
ScreenModuleEditorView "Settings Station Row" 671x200
   TextField "tfLine" at 0,0 size 215x200; Text '$T'
      Visibility <- "Interface.line.visibility"
      Appearance <- "Interface.line.animate"
   TextField "tfLablBtn00" at 215,0 size 40x25; Text '1'
      Visibility <- "Interface.btnRows[0].button.visibility"
      Appearance <- "Interface.btnRows[0].button.animate"
   TextField "tfAllottedBtn00" at 255,0 size 80x25; Text 'Text'
      Visibility <- "Interface.btnRows[0].total.visibility"
      Appearance <- "Interface.btnRows[0].total.animate"
   TextField "tfCriticalBtn00" at 335,0 size 80x25; Text 'Text'
      Visibility <- "Interface.btnRows[0].critical.visibility"
      Appearance <- "Interface.btnRows[0].critical.animate"
   TextField "tfPartNumberBtn00" at 415,0 size 256x25; Text 'Text'
      Visibility <- "Interface.btnRows[0].singlePN.visibility"
      Appearance <- "Interface.btnRows[0].singlePN.animate"
   TextField "tfLablBtn01" at 215,25 size 40x25; Text '2'
      Visibility <- "Interface.btnRows[1].button.visibility"
      Appearance <- "Interface.btnRows[1].button.animate"
   TextField "tfAllottedBtn01" at 255,25 size 80x25; Text 'Text'
      Visibility <- "Interface.btnRows[1].total.visibility"
      Appearance <- "Interface.btnRows[1].total.animate"
   TextField "tfCriticalBtn01" at 335,25 size 80x25; Text 'Text'
      Visibility <- "Interface.btnRows[1].critical.visibility"
      Appearance <- "Interface.btnRows[1].critical.animate"
   TextField "tfPartNumberBtn01" at 415,25 size 256x25; Text 'Text'
      Visibility <- "Interface.btnRows[1].singlePN.visibility"
      Appearance <- "Interface.btnRows[1].singlePN.animate"
   TextField "tfLablBtn02" at 215,50 size 40x25; Text '3'
      Visibility <- "Interface.btnRows[2].button.visibility"
      Appearance <- "Interface.btnRows[2].button.animate"
   TextField "tfAllottedBtn02" at 255,50 size 80x25; Text 'Text'
      Visibility <- "Interface.btnRows[2].total.visibility"
      Appearance <- "Interface.btnRows[2].total.animate"
   TextField "tfCriticalBtn02" at 335,50 size 80x25; Text 'Text'
      Visibility <- "Interface.btnRows[2].critical.visibility"
      Appearance <- "Interface.btnRows[2].critical.animate"
   TextField "tfPartNumberBtn02" at 415,50 size 256x25; Text 'Text'
      Visibility <- "Interface.btnRows[2].singlePN.visibility"
      Appearance <- "Interface.btnRows[2].singlePN.animate"
   TextField "tfLablBtn03" at 215,75 size 40x25; Text '4'
      Visibility <- "Interface.btnRows[3].button.visibility"
      Appearance <- "Interface.btnRows[3].button.animate"
   TextField "tfAllottedBtn03" at 255,75 size 80x25; Text 'Text'
      Visibility <- "Interface.btnRows[3].total.visibility"
      Appearance <- "Interface.btnRows[3].total.animate"
   TextField "tfCriticalBtn03" at 335,75 size 80x25; Text 'Text'
      Visibility <- "Interface.btnRows[3].critical.visibility"
      Appearance <- "Interface.btnRows[3].critical.animate"
   TextField "tfPartNumberBtn03" at 415,75 size 256x25; Text 'Text'
      Visibility <- "Interface.btnRows[3].singlePN.visibility"
      Appearance <- "Interface.btnRows[3].singlePN.animate"
   TextField "tfLablBtn04" at 215,100 size 40x25; Text '5'
      Visibility <- "Interface.btnRows[4].button.visibility"
      Appearance <- "Interface.btnRows[4].button.animate"
   TextField "tfAllottedBtn04" at 255,100 size 80x25; Text 'Text'
      Visibility <- "Interface.btnRows[4].total.visibility"
      Appearance <- "Interface.btnRows[4].total.animate"
   TextField "tfCriticalBtn04" at 335,100 size 80x25; Text 'Text'
      Visibility <- "Interface.btnRows[4].critical.visibility"
      Appearance <- "Interface.btnRows[4].critical.animate"
   TextField "tfPartNumberBtn04" at 415,100 size 256x25; Text 'Text'
      Visibility <- "Interface.btnRows[4].singlePN.visibility"
      Appearance <- "Interface.btnRows[4].singlePN.animate"
   TextField "tfLablBtn05" at 215,125 size 40x25; Text '6'
      Visibility <- "Interface.btnRows[5].button.visibility"
      Appearance <- "Interface.btnRows[5].button.animate"
   TextField "tfAllottedBtn05" at 255,125 size 80x25; Text 'Text'
      Visibility <- "Interface.btnRows[5].total.visibility"
      Appearance <- "Interface.btnRows[5].total.animate"
   TextField "tfCriticalBtn05" at 335,125 size 80x25; Text 'Text'
      Visibility <- "Interface.btnRows[5].critical.visibility"
      Appearance <- "Interface.btnRows[5].critical.animate"
   TextField "tfPartNumberBtn05" at 415,125 size 256x25; Text 'Text'
      Visibility <- "Interface.btnRows[5].singlePN.visibility"
      Appearance <- "Interface.btnRows[5].singlePN.animate"
   TextField "tfLablBtn06" at 215,150 size 40x25; Text '7'
      Visibility <- "Interface.btnRows[6].button.visibility"
      Appearance <- "Interface.btnRows[6].button.animate"
   TextField "tfAllottedBtn06" at 255,150 size 80x25; Text 'Text'
      Visibility <- "Interface.btnRows[6].total.visibility"
      Appearance <- "Interface.btnRows[6].total.animate"
   TextField "tfCriticalBtn06" at 335,150 size 80x25; Text 'Text'
      Visibility <- "Interface.btnRows[6].critical.visibility"
      Appearance <- "Interface.btnRows[6].critical.animate"
   TextField "tfPartNumberBtn06" at 415,150 size 256x25; Text 'Text'
      Visibility <- "Interface.btnRows[6].singlePN.visibility"
      Appearance <- "Interface.btnRows[6].singlePN.animate"
   TextField "tfLablBtn07" at 215,175 size 40x25; Text '8'
      Visibility <- "Interface.btnRows[7].button.visibility"
      Appearance <- "Interface.btnRows[7].button.animate"
   TextField "tfAllottedBtn07" at 255,175 size 80x25; Text 'Text'
      Visibility <- "Interface.btnRows[7].total.visibility"
      Appearance <- "Interface.btnRows[7].total.animate"
   TextField "tfCriticalBtn07" at 335,175 size 80x25; Text 'Text'
      Visibility <- "Interface.btnRows[7].critical.visibility"
      Appearance <- "Interface.btnRows[7].critical.animate"
   TextField "tfPartNumberBtn07" at 415,175 size 256x25; Text 'Text'
      Visibility <- "Interface.btnRows[7].singlePN.visibility"
      Appearance <- "Interface.btnRows[7].singlePN.animate"
   TextField "tfPNDoubleBtn00" at 415,0 size 256x25; Text 'Text'
      Visibility <- "Interface.btnRows[0].doublePN.visibility"
      Appearance <- "Interface.btnRows[0].doublePN.animate"
   TextField "tfPNDoubleBtn01" at 415,25 size 256x25; Text 'Text'
      Visibility <- "Interface.btnRows[1].doublePN.visibility"
      Appearance <- "Interface.btnRows[1].doublePN.animate"
   TextField "tfPNDoubleBtn02" at 415,50 size 256x25; Text 'Text'
      Visibility <- "Interface.btnRows[2].doublePN.visibility"
      Appearance <- "Interface.btnRows[2].doublePN.animate"
   TextField "tfPNDoubleBtn03" at 415,75 size 256x25; Text 'Text'
      Visibility <- "Interface.btnRows[3].doublePN.visibility"
      Appearance <- "Interface.btnRows[3].doublePN.animate"
   TextField "tfPNDoubleBtn04" at 415,100 size 256x25; Text 'Text'
      Visibility <- "Interface.btnRows[4].doublePN.visibility"
      Appearance <- "Interface.btnRows[4].doublePN.animate"
   TextField "tfPNDoubleBtn05" at 415,125 size 256x25; Text 'Text'
      Visibility <- "Interface.btnRows[5].doublePN.visibility"
      Appearance <- "Interface.btnRows[5].doublePN.animate"
   TextField "tfPNDoubleBtn06" at 415,150 size 256x25; Text 'Text'
      Visibility <- "Interface.btnRows[6].doublePN.visibility"
      Appearance <- "Interface.btnRows[6].doublePN.animate"
   TextField "tfPNDoubleBtn07" at 415,175 size 256x25; Text 'Text'
      Visibility <- "Interface.btnRows[7].doublePN.visibility"
      Appearance <- "Interface.btnRows[7].doublePN.animate"
*)

(* ===== HMI "HMI_RT_1" =====

ScreenModuleEditorView "Settings Station Row" 671x200
   TextField "tfLine" at 0,0 size 215x200; Text 'Text'
      Visibility <- "Interface.line.visibility"
      Appearance <- "Interface.line.animate"
   TextField "tfLablBtn00" at 215,0 size 40x25; Text '1'
      Visibility <- "Interface.btnRows[0].button.visibility"
      Appearance <- "Interface.btnRows[0].button.animate"
   TextField "tfAllottedBtn00" at 255,0 size 80x25; Text 'Text'
      Visibility <- "Interface.btnRows[0].total.visibility"
      Appearance <- "Interface.btnRows[0].total.animate"
   TextField "tfCriticalBtn00" at 335,0 size 80x25; Text 'Text'
      Visibility <- "Interface.btnRows[0].critical.visibility"
      Appearance <- "Interface.btnRows[0].critical.animate"
   TextField "tfPartNumberBtn00" at 415,0 size 256x25; Text 'Text'
      Visibility <- "Interface.btnRows[0].singlePN.visibility"
      Appearance <- "Interface.btnRows[0].singlePN.animate"
   TextField "tfLablBtn01" at 215,25 size 40x25; Text '2'
      Visibility <- "Interface.btnRows[1].button.visibility"
      Appearance <- "Interface.btnRows[1].button.animate"
   TextField "tfAllottedBtn01" at 255,25 size 80x25; Text 'Text'
      Visibility <- "Interface.btnRows[1].total.visibility"
      Appearance <- "Interface.btnRows[1].total.animate"
   TextField "tfCriticalBtn01" at 335,25 size 80x25; Text 'Text'
      Visibility <- "Interface.btnRows[1].critical.visibility"
      Appearance <- "Interface.btnRows[1].critical.animate"
   TextField "tfPartNumberBtn01" at 415,25 size 256x25; Text 'Text'
      Visibility <- "Interface.btnRows[1].singlePN.visibility"
      Appearance <- "Interface.btnRows[1].singlePN.animate"
   TextField "tfLablBtn02" at 215,50 size 40x25; Text '3'
      Visibility <- "Interface.btnRows[2].button.visibility"
      Appearance <- "Interface.btnRows[2].button.animate"
   TextField "tfAllottedBtn02" at 255,50 size 80x25; Text 'Text'
      Visibility <- "Interface.btnRows[2].total.visibility"
      Appearance <- "Interface.btnRows[2].total.animate"
   TextField "tfCriticalBtn02" at 335,50 size 80x25; Text 'Text'
      Visibility <- "Interface.btnRows[2].critical.visibility"
      Appearance <- "Interface.btnRows[2].critical.animate"
   TextField "tfPartNumberBtn02" at 415,50 size 256x25; Text 'Text'
      Visibility <- "Interface.btnRows[2].singlePN.visibility"
      Appearance <- "Interface.btnRows[2].singlePN.animate"
   TextField "tfLablBtn03" at 215,75 size 40x25; Text '4'
      Visibility <- "Interface.btnRows[3].button.visibility"
      Appearance <- "Interface.btnRows[3].button.animate"
   TextField "tfAllottedBtn03" at 255,75 size 80x25; Text 'Text'
      Visibility <- "Interface.btnRows[3].total.visibility"
      Appearance <- "Interface.btnRows[3].total.animate"
   TextField "tfCriticalBtn03" at 335,75 size 80x25; Text 'Text'
      Visibility <- "Interface.btnRows[3].critical.visibility"
      Appearance <- "Interface.btnRows[3].critical.animate"
   TextField "tfPartNumberBtn03" at 415,75 size 256x25; Text 'Text'
      Visibility <- "Interface.btnRows[3].singlePN.visibility"
      Appearance <- "Interface.btnRows[3].singlePN.animate"
   TextField "tfLablBtn04" at 215,100 size 40x25; Text '5'
      Visibility <- "Interface.btnRows[4].button.visibility"
      Appearance <- "Interface.btnRows[4].button.animate"
   TextField "tfAllottedBtn04" at 255,100 size 80x25; Text 'Text'
      Visibility <- "Interface.btnRows[4].total.visibility"
      Appearance <- "Interface.btnRows[4].total.animate"
   TextField "tfCriticalBtn04" at 335,100 size 80x25; Text 'Text'
      Visibility <- "Interface.btnRows[4].critical.visibility"
      Appearance <- "Interface.btnRows[4].critical.animate"
   TextField "tfPartNumberBtn04" at 415,100 size 256x25; Text 'Text'
      Visibility <- "Interface.btnRows[4].singlePN.visibility"
      Appearance <- "Interface.btnRows[4].singlePN.animate"
   TextField "tfLablBtn05" at 215,125 size 40x25; Text '6'
      Visibility <- "Interface.btnRows[5].button.visibility"
      Appearance <- "Interface.btnRows[5].button.animate"
   TextField "tfAllottedBtn05" at 255,125 size 80x25; Text 'Text'
      Visibility <- "Interface.btnRows[5].total.visibility"
      Appearance <- "Interface.btnRows[5].total.animate"
   TextField "tfCriticalBtn05" at 335,125 size 80x25; Text 'Text'
      Visibility <- "Interface.btnRows[5].critical.visibility"
      Appearance <- "Interface.btnRows[5].critical.animate"
   TextField "tfPartNumberBtn05" at 415,125 size 256x25; Text 'Text'
      Visibility <- "Interface.btnRows[5].singlePN.visibility"
      Appearance <- "Interface.btnRows[5].singlePN.animate"
   TextField "tfLablBtn06" at 215,150 size 40x25; Text '7'
      Visibility <- "Interface.btnRows[6].button.visibility"
      Appearance <- "Interface.btnRows[6].button.animate"
   TextField "tfAllottedBtn06" at 255,150 size 80x25; Text 'Text'
      Visibility <- "Interface.btnRows[6].total.visibility"
      Appearance <- "Interface.btnRows[6].total.animate"
   TextField "tfCriticalBtn06" at 335,150 size 80x25; Text 'Text'
      Visibility <- "Interface.btnRows[6].critical.visibility"
      Appearance <- "Interface.btnRows[6].critical.animate"
   TextField "tfPartNumberBtn06" at 415,150 size 256x25; Text 'Text'
      Visibility <- "Interface.btnRows[6].singlePN.visibility"
      Appearance <- "Interface.btnRows[6].singlePN.animate"
   TextField "tfLablBtn07" at 215,175 size 40x25; Text '8'
      Visibility <- "Interface.btnRows[7].button.visibility"
      Appearance <- "Interface.btnRows[7].button.animate"
   TextField "tfAllottedBtn07" at 255,175 size 80x25; Text 'Text'
      Visibility <- "Interface.btnRows[7].total.visibility"
      Appearance <- "Interface.btnRows[7].total.animate"
   TextField "tfCriticalBtn07" at 335,175 size 80x25; Text 'Text'
      Visibility <- "Interface.btnRows[7].critical.visibility"
      Appearance <- "Interface.btnRows[7].critical.animate"
   TextField "tfPartNumberBtn07" at 415,175 size 256x25; Text 'Text'
      Visibility <- "Interface.btnRows[7].singlePN.visibility"
      Appearance <- "Interface.btnRows[7].singlePN.animate"
   TextField "tfPNDoubleBtn00" at 415,0 size 256x25; Text 'Text'
      Visibility <- "Interface.btnRows[0].doublePN.visibility"
      Appearance <- "Interface.btnRows[0].doublePN.animate"
   TextField "tfPNDoubleBtn01" at 415,25 size 256x25; Text 'Text'
      Visibility <- "Interface.btnRows[1].doublePN.visibility"
      Appearance <- "Interface.btnRows[1].doublePN.animate"
   TextField "tfPNDoubleBtn02" at 415,50 size 256x25; Text 'Text'
      Visibility <- "Interface.btnRows[2].doublePN.visibility"
      Appearance <- "Interface.btnRows[2].doublePN.animate"
   TextField "tfPNDoubleBtn03" at 415,75 size 256x25; Text 'Text'
      Visibility <- "Interface.btnRows[3].doublePN.visibility"
      Appearance <- "Interface.btnRows[3].doublePN.animate"
   TextField "tfPNDoubleBtn04" at 415,100 size 256x25; Text 'Text'
      Visibility <- "Interface.btnRows[4].doublePN.visibility"
      Appearance <- "Interface.btnRows[4].doublePN.animate"
   TextField "tfPNDoubleBtn05" at 415,125 size 256x25; Text 'Text'
      Visibility <- "Interface.btnRows[5].doublePN.visibility"
      Appearance <- "Interface.btnRows[5].doublePN.animate"
   TextField "tfPNDoubleBtn06" at 415,150 size 256x25; Text 'Text'
      Visibility <- "Interface.btnRows[6].doublePN.visibility"
      Appearance <- "Interface.btnRows[6].doublePN.animate"
   TextField "tfPNDoubleBtn07" at 415,175 size 256x25; Text 'Text'
      Visibility <- "Interface.btnRows[7].doublePN.visibility"
      Appearance <- "Interface.btnRows[7].doublePN.animate"
*)

(* ===== HMI "HMI_RT_1" =====

ScreenModuleEditorView "Settings Station Row" 671x200
   TextField "tfLine" at 0,0 size 215x200; Text 'Text'
      Visibility <- "Interface.line.visibility"
      Appearance <- "Interface.line.animate"
   TextField "tfLablBtn00" at 215,0 size 40x25; Text '1'
      Visibility <- "Interface.btnRows[0].button.visibility"
      Appearance <- "Interface.btnRows[0].button.animate"
   TextField "tfAllottedBtn00" at 255,0 size 80x25; Text 'Text'
      Visibility <- "Interface.btnRows[0].total.visibility"
      Appearance <- "Interface.btnRows[0].total.animate"
   TextField "tfCriticalBtn00" at 335,0 size 80x25; Text 'Text'
      Visibility <- "Interface.btnRows[0].critical.visibility"
      Appearance <- "Interface.btnRows[0].critical.animate"
   TextField "tfPartNumberBtn00" at 415,0 size 256x25; Text 'Text'
      Visibility <- "Interface.btnRows[0].singlePN.visibility"
      Appearance <- "Interface.btnRows[0].singlePN.animate"
   TextField "tfLablBtn01" at 215,25 size 40x25; Text '2'
      Visibility <- "Interface.btnRows[1].button.visibility"
      Appearance <- "Interface.btnRows[1].button.animate"
   TextField "tfAllottedBtn01" at 255,25 size 80x25; Text 'Text'
      Visibility <- "Interface.btnRows[1].total.visibility"
      Appearance <- "Interface.btnRows[1].total.animate"
   TextField "tfCriticalBtn01" at 335,25 size 80x25; Text 'Text'
      Visibility <- "Interface.btnRows[1].critical.visibility"
      Appearance <- "Interface.btnRows[1].critical.animate"
   TextField "tfPartNumberBtn01" at 415,25 size 256x25; Text 'Text'
      Visibility <- "Interface.btnRows[1].singlePN.visibility"
      Appearance <- "Interface.btnRows[1].singlePN.animate"
   TextField "tfLablBtn02" at 215,50 size 40x25; Text '3'
      Visibility <- "Interface.btnRows[2].button.visibility"
      Appearance <- "Interface.btnRows[2].button.animate"
   TextField "tfAllottedBtn02" at 255,50 size 80x25; Text 'Text'
      Visibility <- "Interface.btnRows[2].total.visibility"
      Appearance <- "Interface.btnRows[2].total.animate"
   TextField "tfCriticalBtn02" at 335,50 size 80x25; Text 'Text'
      Visibility <- "Interface.btnRows[2].critical.visibility"
      Appearance <- "Interface.btnRows[2].critical.animate"
   TextField "tfPartNumberBtn02" at 415,50 size 256x25; Text 'Text'
      Visibility <- "Interface.btnRows[2].singlePN.visibility"
      Appearance <- "Interface.btnRows[2].singlePN.animate"
   TextField "tfLablBtn03" at 215,75 size 40x25; Text '4'
      Visibility <- "Interface.btnRows[3].button.visibility"
      Appearance <- "Interface.btnRows[3].button.animate"
   TextField "tfAllottedBtn03" at 255,75 size 80x25; Text 'Text'
      Visibility <- "Interface.btnRows[3].total.visibility"
      Appearance <- "Interface.btnRows[3].total.animate"
   TextField "tfCriticalBtn03" at 335,75 size 80x25; Text 'Text'
      Visibility <- "Interface.btnRows[3].critical.visibility"
      Appearance <- "Interface.btnRows[3].critical.animate"
   TextField "tfPartNumberBtn03" at 415,75 size 256x25; Text 'Text'
      Visibility <- "Interface.btnRows[3].singlePN.visibility"
      Appearance <- "Interface.btnRows[3].singlePN.animate"
   TextField "tfLablBtn04" at 215,100 size 40x25; Text '5'
      Visibility <- "Interface.btnRows[4].button.visibility"
      Appearance <- "Interface.btnRows[4].button.animate"
   TextField "tfAllottedBtn04" at 255,100 size 80x25; Text 'Text'
      Visibility <- "Interface.btnRows[4].total.visibility"
      Appearance <- "Interface.btnRows[4].total.animate"
   TextField "tfCriticalBtn04" at 335,100 size 80x25; Text 'Text'
      Visibility <- "Interface.btnRows[4].critical.visibility"
      Appearance <- "Interface.btnRows[4].critical.animate"
   TextField "tfPartNumberBtn04" at 415,100 size 256x25; Text 'Text'
      Visibility <- "Interface.btnRows[4].singlePN.visibility"
      Appearance <- "Interface.btnRows[4].singlePN.animate"
   TextField "tfLablBtn05" at 215,125 size 40x25; Text '6'
      Visibility <- "Interface.btnRows[5].button.visibility"
      Appearance <- "Interface.btnRows[5].button.animate"
   TextField "tfAllottedBtn05" at 255,125 size 80x25; Text 'Text'
      Visibility <- "Interface.btnRows[5].total.visibility"
      Appearance <- "Interface.btnRows[5].total.animate"
   TextField "tfCriticalBtn05" at 335,125 size 80x25; Text 'Text'
      Visibility <- "Interface.btnRows[5].critical.visibility"
      Appearance <- "Interface.btnRows[5].critical.animate"
   TextField "tfPartNumberBtn05" at 415,125 size 256x25; Text 'Text'
      Visibility <- "Interface.btnRows[5].singlePN.visibility"
      Appearance <- "Interface.btnRows[5].singlePN.animate"
   TextField "tfLablBtn06" at 215,150 size 40x25; Text '7'
      Visibility <- "Interface.btnRows[6].button.visibility"
      Appearance <- "Interface.btnRows[6].button.animate"
   TextField "tfAllottedBtn06" at 255,150 size 80x25; Text 'Text'
      Visibility <- "Interface.btnRows[6].total.visibility"
      Appearance <- "Interface.btnRows[6].total.animate"
   TextField "tfCriticalBtn06" at 335,150 size 80x25; Text 'Text'
      Visibility <- "Interface.btnRows[6].critical.visibility"
      Appearance <- "Interface.btnRows[6].critical.animate"
   TextField "tfPartNumberBtn06" at 415,150 size 256x25; Text 'Text'
      Visibility <- "Interface.btnRows[6].singlePN.visibility"
      Appearance <- "Interface.btnRows[6].singlePN.animate"
   TextField "tfLablBtn07" at 215,175 size 40x25; Text '8'
      Visibility <- "Interface.btnRows[7].button.visibility"
      Appearance <- "Interface.btnRows[7].button.animate"
   TextField "tfAllottedBtn07" at 255,175 size 80x25; Text 'Text'
      Visibility <- "Interface.btnRows[7].total.visibility"
      Appearance <- "Interface.btnRows[7].total.animate"
   TextField "tfCriticalBtn07" at 335,175 size 80x25; Text 'Text'
      Visibility <- "Interface.btnRows[7].critical.visibility"
      Appearance <- "Interface.btnRows[7].critical.animate"
   TextField "tfPartNumberBtn07" at 415,175 size 256x25; Text 'Text'
      Visibility <- "Interface.btnRows[7].singlePN.visibility"
      Appearance <- "Interface.btnRows[7].singlePN.animate"
   TextField "tfPNDoubleBtn00" at 415,0 size 256x25; Text 'Text'
      Visibility <- "Interface.btnRows[0].doublePN.visibility"
      Appearance <- "Interface.btnRows[0].doublePN.animate"
   TextField "tfPNDoubleBtn01" at 415,25 size 256x25; Text 'Text'
      Visibility <- "Interface.btnRows[1].doublePN.visibility"
      Appearance <- "Interface.btnRows[1].doublePN.animate"
   TextField "tfPNDoubleBtn02" at 415,50 size 256x25; Text 'Text'
      Visibility <- "Interface.btnRows[2].doublePN.visibility"
      Appearance <- "Interface.btnRows[2].doublePN.animate"
   TextField "tfPNDoubleBtn03" at 415,75 size 256x25; Text 'Text'
      Visibility <- "Interface.btnRows[3].doublePN.visibility"
      Appearance <- "Interface.btnRows[3].doublePN.animate"
   TextField "tfPNDoubleBtn04" at 415,100 size 256x25; Text 'Text'
      Visibility <- "Interface.btnRows[4].doublePN.visibility"
      Appearance <- "Interface.btnRows[4].doublePN.animate"
   TextField "tfPNDoubleBtn05" at 415,125 size 256x25; Text 'Text'
      Visibility <- "Interface.btnRows[5].doublePN.visibility"
      Appearance <- "Interface.btnRows[5].doublePN.animate"
   TextField "tfPNDoubleBtn06" at 415,150 size 256x25; Text 'Text'
      Visibility <- "Interface.btnRows[6].doublePN.visibility"
      Appearance <- "Interface.btnRows[6].doublePN.animate"
   TextField "tfPNDoubleBtn07" at 415,175 size 256x25; Text 'Text'
      Visibility <- "Interface.btnRows[7].doublePN.visibility"
      Appearance <- "Interface.btnRows[7].doublePN.animate"
*)

(* ===== HMI "HMI_RT_1" =====

ScreenModuleEditorView "Settings Station Row" 671x200
   TextField "tfLine" at 0,0 size 215x200; Text 'Text'
      Visibility <- "Interface.line.visibility"
      Appearance <- "Interface.line.animate"
   TextField "tfLablBtn00" at 215,0 size 40x25; Text '1'
      Visibility <- "Interface.btnRows[0].button.visibility"
      Appearance <- "Interface.btnRows[0].button.animate"
   TextField "tfAllottedBtn00" at 255,0 size 80x25; Text 'Text'
      Visibility <- "Interface.btnRows[0].total.visibility"
      Appearance <- "Interface.btnRows[0].total.animate"
   TextField "tfCriticalBtn00" at 335,0 size 80x25; Text 'Text'
      Visibility <- "Interface.btnRows[0].critical.visibility"
      Appearance <- "Interface.btnRows[0].critical.animate"
   TextField "tfPartNumberBtn00" at 415,0 size 256x25; Text 'Text'
      Visibility <- "Interface.btnRows[0].singlePN.visibility"
      Appearance <- "Interface.btnRows[0].singlePN.animate"
   TextField "tfLablBtn01" at 215,25 size 40x25; Text '2'
      Visibility <- "Interface.btnRows[1].button.visibility"
      Appearance <- "Interface.btnRows[1].button.animate"
   TextField "tfAllottedBtn01" at 255,25 size 80x25; Text 'Text'
      Visibility <- "Interface.btnRows[1].total.visibility"
      Appearance <- "Interface.btnRows[1].total.animate"
   TextField "tfCriticalBtn01" at 335,25 size 80x25; Text 'Text'
      Visibility <- "Interface.btnRows[1].critical.visibility"
      Appearance <- "Interface.btnRows[1].critical.animate"
   TextField "tfPartNumberBtn01" at 415,25 size 256x25; Text 'Text'
      Visibility <- "Interface.btnRows[1].singlePN.visibility"
      Appearance <- "Interface.btnRows[1].singlePN.animate"
   TextField "tfLablBtn02" at 215,50 size 40x25; Text '3'
      Visibility <- "Interface.btnRows[2].button.visibility"
      Appearance <- "Interface.btnRows[2].button.animate"
   TextField "tfAllottedBtn02" at 255,50 size 80x25; Text 'Text'
      Visibility <- "Interface.btnRows[2].total.visibility"
      Appearance <- "Interface.btnRows[2].total.animate"
   TextField "tfCriticalBtn02" at 335,50 size 80x25; Text 'Text'
      Visibility <- "Interface.btnRows[2].critical.visibility"
      Appearance <- "Interface.btnRows[2].critical.animate"
   TextField "tfPartNumberBtn02" at 415,50 size 256x25; Text 'Text'
      Visibility <- "Interface.btnRows[2].singlePN.visibility"
      Appearance <- "Interface.btnRows[2].singlePN.animate"
   TextField "tfLablBtn03" at 215,75 size 40x25; Text '4'
      Visibility <- "Interface.btnRows[3].button.visibility"
      Appearance <- "Interface.btnRows[3].button.animate"
   TextField "tfAllottedBtn03" at 255,75 size 80x25; Text 'Text'
      Visibility <- "Interface.btnRows[3].total.visibility"
      Appearance <- "Interface.btnRows[3].total.animate"
   TextField "tfCriticalBtn03" at 335,75 size 80x25; Text 'Text'
      Visibility <- "Interface.btnRows[3].critical.visibility"
      Appearance <- "Interface.btnRows[3].critical.animate"
   TextField "tfPartNumberBtn03" at 415,75 size 256x25; Text 'Text'
      Visibility <- "Interface.btnRows[3].singlePN.visibility"
      Appearance <- "Interface.btnRows[3].singlePN.animate"
   TextField "tfLablBtn04" at 215,100 size 40x25; Text '5'
      Visibility <- "Interface.btnRows[4].button.visibility"
      Appearance <- "Interface.btnRows[4].button.animate"
   TextField "tfAllottedBtn04" at 255,100 size 80x25; Text 'Text'
      Visibility <- "Interface.btnRows[4].total.visibility"
      Appearance <- "Interface.btnRows[4].total.animate"
   TextField "tfCriticalBtn04" at 335,100 size 80x25; Text 'Text'
      Visibility <- "Interface.btnRows[4].critical.visibility"
      Appearance <- "Interface.btnRows[4].critical.animate"
   TextField "tfPartNumberBtn04" at 415,100 size 256x25; Text 'Text'
      Visibility <- "Interface.btnRows[4].singlePN.visibility"
      Appearance <- "Interface.btnRows[4].singlePN.animate"
   TextField "tfLablBtn05" at 215,125 size 40x25; Text '6'
      Visibility <- "Interface.btnRows[5].button.visibility"
      Appearance <- "Interface.btnRows[5].button.animate"
   TextField "tfAllottedBtn05" at 255,125 size 80x25; Text 'Text'
      Visibility <- "Interface.btnRows[5].total.visibility"
      Appearance <- "Interface.btnRows[5].total.animate"
   TextField "tfCriticalBtn05" at 335,125 size 80x25; Text 'Text'
      Visibility <- "Interface.btnRows[5].critical.visibility"
      Appearance <- "Interface.btnRows[5].critical.animate"
   TextField "tfPartNumberBtn05" at 415,125 size 256x25; Text 'Text'
      Visibility <- "Interface.btnRows[5].singlePN.visibility"
      Appearance <- "Interface.btnRows[5].singlePN.animate"
   TextField "tfLablBtn06" at 215,150 size 40x25; Text '7'
      Visibility <- "Interface.btnRows[6].button.visibility"
      Appearance <- "Interface.btnRows[6].button.animate"
   TextField "tfAllottedBtn06" at 255,150 size 80x25; Text 'Text'
      Visibility <- "Interface.btnRows[6].total.visibility"
      Appearance <- "Interface.btnRows[6].total.animate"
   TextField "tfCriticalBtn06" at 335,150 size 80x25; Text 'Text'
      Visibility <- "Interface.btnRows[6].critical.visibility"
      Appearance <- "Interface.btnRows[6].critical.animate"
   TextField "tfPartNumberBtn06" at 415,150 size 256x25; Text 'Text'
      Visibility <- "Interface.btnRows[6].singlePN.visibility"
      Appearance <- "Interface.btnRows[6].singlePN.animate"
   TextField "tfLablBtn07" at 215,175 size 40x25; Text '8'
      Visibility <- "Interface.btnRows[7].button.visibility"
      Appearance <- "Interface.btnRows[7].button.animate"
   TextField "tfAllottedBtn07" at 255,175 size 80x25; Text 'Text'
      Visibility <- "Interface.btnRows[7].total.visibility"
      Appearance <- "Interface.btnRows[7].total.animate"
   TextField "tfCriticalBtn07" at 335,175 size 80x25; Text 'Text'
      Visibility <- "Interface.btnRows[7].critical.visibility"
      Appearance <- "Interface.btnRows[7].critical.animate"
   TextField "tfPartNumberBtn07" at 415,175 size 256x25; Text 'Text'
      Visibility <- "Interface.btnRows[7].singlePN.visibility"
      Appearance <- "Interface.btnRows[7].singlePN.animate"
   TextField "tfPNDoubleBtn00" at 415,0 size 256x25; Text 'Text'
      Visibility <- "Interface.btnRows[0].doublePN.visibility"
      Appearance <- "Interface.btnRows[0].doublePN.animate"
   TextField "tfPNDoubleBtn01" at 415,25 size 256x25; Text 'Text'
      Visibility <- "Interface.btnRows[1].doublePN.visibility"
      Appearance <- "Interface.btnRows[1].doublePN.animate"
   TextField "tfPNDoubleBtn02" at 415,50 size 256x25; Text 'Text'
      Visibility <- "Interface.btnRows[2].doublePN.visibility"
      Appearance <- "Interface.btnRows[2].doublePN.animate"
   TextField "tfPNDoubleBtn03" at 415,75 size 256x25; Text 'Text'
      Visibility <- "Interface.btnRows[3].doublePN.visibility"
      Appearance <- "Interface.btnRows[3].doublePN.animate"
   TextField "tfPNDoubleBtn04" at 415,100 size 256x25; Text 'Text'
      Visibility <- "Interface.btnRows[4].doublePN.visibility"
      Appearance <- "Interface.btnRows[4].doublePN.animate"
   TextField "tfPNDoubleBtn05" at 415,125 size 256x25; Text 'Text'
      Visibility <- "Interface.btnRows[5].doublePN.visibility"
      Appearance <- "Interface.btnRows[5].doublePN.animate"
   TextField "tfPNDoubleBtn06" at 415,150 size 256x25; Text 'Text'
      Visibility <- "Interface.btnRows[6].doublePN.visibility"
      Appearance <- "Interface.btnRows[6].doublePN.animate"
   TextField "tfPNDoubleBtn07" at 415,175 size 256x25; Text 'Text'
      Visibility <- "Interface.btnRows[7].doublePN.visibility"
      Appearance <- "Interface.btnRows[7].doublePN.animate"
*)

(* ===== HMI "HMI_RT_1" =====

ScreenModuleEditorView "Settings Station Row" 671x200
   TextField "tfLine" at 0,0 size 215x200; Text 'Text'
      Visibility <- "Interface.line.visibility"
      Appearance <- "Interface.line.animate"
   TextField "tfLablBtn00" at 215,0 size 40x25; Text '1'
      Visibility <- "Interface.btnRows[0].button.visibility"
      Appearance <- "Interface.btnRows[0].button.animate"
   TextField "tfAllottedBtn00" at 255,0 size 80x25; Text 'Text'
      Visibility <- "Interface.btnRows[0].total.visibility"
      Appearance <- "Interface.btnRows[0].total.animate"
   TextField "tfCriticalBtn00" at 335,0 size 80x25; Text 'Text'
      Visibility <- "Interface.btnRows[0].critical.visibility"
      Appearance <- "Interface.btnRows[0].critical.animate"
   TextField "tfPartNumberBtn00" at 415,0 size 256x25; Text 'Text'
      Visibility <- "Interface.btnRows[0].singlePN.visibility"
      Appearance <- "Interface.btnRows[0].singlePN.animate"
   TextField "tfLablBtn01" at 215,25 size 40x25; Text '2'
      Visibility <- "Interface.btnRows[1].button.visibility"
      Appearance <- "Interface.btnRows[1].button.animate"
   TextField "tfAllottedBtn01" at 255,25 size 80x25; Text 'Text'
      Visibility <- "Interface.btnRows[1].total.visibility"
      Appearance <- "Interface.btnRows[1].total.animate"
   TextField "tfCriticalBtn01" at 335,25 size 80x25; Text 'Text'
      Visibility <- "Interface.btnRows[1].critical.visibility"
      Appearance <- "Interface.btnRows[1].critical.animate"
   TextField "tfPartNumberBtn01" at 415,25 size 256x25; Text 'Text'
      Visibility <- "Interface.btnRows[1].singlePN.visibility"
      Appearance <- "Interface.btnRows[1].singlePN.animate"
   TextField "tfLablBtn02" at 215,50 size 40x25; Text '3'
      Visibility <- "Interface.btnRows[2].button.visibility"
      Appearance <- "Interface.btnRows[2].button.animate"
   TextField "tfAllottedBtn02" at 255,50 size 80x25; Text 'Text'
      Visibility <- "Interface.btnRows[2].total.visibility"
      Appearance <- "Interface.btnRows[2].total.animate"
   TextField "tfCriticalBtn02" at 335,50 size 80x25; Text 'Text'
      Visibility <- "Interface.btnRows[2].critical.visibility"
      Appearance <- "Interface.btnRows[2].critical.animate"
   TextField "tfPartNumberBtn02" at 415,50 size 256x25; Text 'Text'
      Visibility <- "Interface.btnRows[2].singlePN.visibility"
      Appearance <- "Interface.btnRows[2].singlePN.animate"
   TextField "tfLablBtn03" at 215,75 size 40x25; Text '4'
      Visibility <- "Interface.btnRows[3].button.visibility"
      Appearance <- "Interface.btnRows[3].button.animate"
   TextField "tfAllottedBtn03" at 255,75 size 80x25; Text 'Text'
      Visibility <- "Interface.btnRows[3].total.visibility"
      Appearance <- "Interface.btnRows[3].total.animate"
   TextField "tfCriticalBtn03" at 335,75 size 80x25; Text 'Text'
      Visibility <- "Interface.btnRows[3].critical.visibility"
      Appearance <- "Interface.btnRows[3].critical.animate"
   TextField "tfPartNumberBtn03" at 415,75 size 256x25; Text 'Text'
      Visibility <- "Interface.btnRows[3].singlePN.visibility"
      Appearance <- "Interface.btnRows[3].singlePN.animate"
   TextField "tfLablBtn04" at 215,100 size 40x25; Text '5'
      Visibility <- "Interface.btnRows[4].button.visibility"
      Appearance <- "Interface.btnRows[4].button.animate"
   TextField "tfAllottedBtn04" at 255,100 size 80x25; Text 'Text'
      Visibility <- "Interface.btnRows[4].total.visibility"
      Appearance <- "Interface.btnRows[4].total.animate"
   TextField "tfCriticalBtn04" at 335,100 size 80x25; Text 'Text'
      Visibility <- "Interface.btnRows[4].critical.visibility"
      Appearance <- "Interface.btnRows[4].critical.animate"
   TextField "tfPartNumberBtn04" at 415,100 size 256x25; Text 'Text'
      Visibility <- "Interface.btnRows[4].singlePN.visibility"
      Appearance <- "Interface.btnRows[4].singlePN.animate"
   TextField "tfLablBtn05" at 215,125 size 40x25; Text '6'
      Visibility <- "Interface.btnRows[5].button.visibility"
      Appearance <- "Interface.btnRows[5].button.animate"
   TextField "tfAllottedBtn05" at 255,125 size 80x25; Text 'Text'
      Visibility <- "Interface.btnRows[5].total.visibility"
      Appearance <- "Interface.btnRows[5].total.animate"
   TextField "tfCriticalBtn05" at 335,125 size 80x25; Text 'Text'
      Visibility <- "Interface.btnRows[5].critical.visibility"
      Appearance <- "Interface.btnRows[5].critical.animate"
   TextField "tfPartNumberBtn05" at 415,125 size 256x25; Text 'Text'
      Visibility <- "Interface.btnRows[5].singlePN.visibility"
      Appearance <- "Interface.btnRows[5].singlePN.animate"
   TextField "tfLablBtn06" at 215,150 size 40x25; Text '7'
      Visibility <- "Interface.btnRows[6].button.visibility"
      Appearance <- "Interface.btnRows[6].button.animate"
   TextField "tfAllottedBtn06" at 255,150 size 80x25; Text 'Text'
      Visibility <- "Interface.btnRows[6].total.visibility"
      Appearance <- "Interface.btnRows[6].total.animate"
   TextField "tfCriticalBtn06" at 335,150 size 80x25; Text 'Text'
      Visibility <- "Interface.btnRows[6].critical.visibility"
      Appearance <- "Interface.btnRows[6].critical.animate"
   TextField "tfPartNumberBtn06" at 415,150 size 256x25; Text 'Text'
      Visibility <- "Interface.btnRows[6].singlePN.visibility"
      Appearance <- "Interface.btnRows[6].singlePN.animate"
   TextField "tfLablBtn07" at 215,175 size 40x25; Text '8'
      Visibility <- "Interface.btnRows[7].button.visibility"
      Appearance <- "Interface.btnRows[7].button.animate"
   TextField "tfAllottedBtn07" at 255,175 size 80x25; Text 'Text'
      Visibility <- "Interface.btnRows[7].total.visibility"
      Appearance <- "Interface.btnRows[7].total.animate"
   TextField "tfCriticalBtn07" at 335,175 size 80x25; Text 'Text'
      Visibility <- "Interface.btnRows[7].critical.visibility"
      Appearance <- "Interface.btnRows[7].critical.animate"
   TextField "tfPartNumberBtn07" at 415,175 size 256x25; Text 'Text'
      Visibility <- "Interface.btnRows[7].singlePN.visibility"
      Appearance <- "Interface.btnRows[7].singlePN.animate"
   TextField "tfPNDoubleBtn00" at 415,0 size 256x25; Text 'Text'
      Visibility <- "Interface.btnRows[0].doublePN.visibility"
      Appearance <- "Interface.btnRows[0].doublePN.animate"
   TextField "tfPNDoubleBtn01" at 415,25 size 256x25; Text 'Text'
      Visibility <- "Interface.btnRows[1].doublePN.visibility"
      Appearance <- "Interface.btnRows[1].doublePN.animate"
   TextField "tfPNDoubleBtn02" at 415,50 size 256x25; Text 'Text'
      Visibility <- "Interface.btnRows[2].doublePN.visibility"
      Appearance <- "Interface.btnRows[2].doublePN.animate"
   TextField "tfPNDoubleBtn03" at 415,75 size 256x25; Text 'Text'
      Visibility <- "Interface.btnRows[3].doublePN.visibility"
      Appearance <- "Interface.btnRows[3].doublePN.animate"
   TextField "tfPNDoubleBtn04" at 415,100 size 256x25; Text 'Text'
      Visibility <- "Interface.btnRows[4].doublePN.visibility"
      Appearance <- "Interface.btnRows[4].doublePN.animate"
   TextField "tfPNDoubleBtn05" at 415,125 size 256x25; Text 'Text'
      Visibility <- "Interface.btnRows[5].doublePN.visibility"
      Appearance <- "Interface.btnRows[5].doublePN.animate"
   TextField "tfPNDoubleBtn06" at 415,150 size 256x25; Text 'Text'
      Visibility <- "Interface.btnRows[6].doublePN.visibility"
      Appearance <- "Interface.btnRows[6].doublePN.animate"
   TextField "tfPNDoubleBtn07" at 415,175 size 256x25; Text 'Text'
      Visibility <- "Interface.btnRows[7].doublePN.visibility"
      Appearance <- "Interface.btnRows[7].doublePN.animate"
*)

(* ===== HMI "HMI_RT_1" =====

ScreenModuleEditorView "Settings Station Row" 671x200
   TextField "tfLine" at 0,0 size 215x200; Text 'Text'
      Visibility <- "Interface.line.visibility"
      Appearance <- "Interface.line.animate"
   TextField "tfLablBtn00" at 215,0 size 40x25; Text '1'
      Visibility <- "Interface.btnRows[0].button.visibility"
      Appearance <- "Interface.btnRows[0].button.animate"
   TextField "tfAllottedBtn00" at 255,0 size 80x25; Text 'Text'
      Visibility <- "Interface.btnRows[0].total.visibility"
      Appearance <- "Interface.btnRows[0].total.animate"
   TextField "tfCriticalBtn00" at 335,0 size 80x25; Text 'Text'
      Visibility <- "Interface.btnRows[0].critical.visibility"
      Appearance <- "Interface.btnRows[0].critical.animate"
   TextField "tfPartNumberBtn00" at 415,0 size 256x25; Text 'Text'
      Visibility <- "Interface.btnRows[0].singlePN.visibility"
      Appearance <- "Interface.btnRows[0].singlePN.animate"
   TextField "tfLablBtn01" at 215,25 size 40x25; Text '2'
      Visibility <- "Interface.btnRows[1].button.visibility"
      Appearance <- "Interface.btnRows[1].button.animate"
   TextField "tfAllottedBtn01" at 255,25 size 80x25; Text 'Text'
      Visibility <- "Interface.btnRows[1].total.visibility"
      Appearance <- "Interface.btnRows[1].total.animate"
   TextField "tfCriticalBtn01" at 335,25 size 80x25; Text 'Text'
      Visibility <- "Interface.btnRows[1].critical.visibility"
      Appearance <- "Interface.btnRows[1].critical.animate"
   TextField "tfPartNumberBtn01" at 415,25 size 256x25; Text 'Text'
      Visibility <- "Interface.btnRows[1].singlePN.visibility"
      Appearance <- "Interface.btnRows[1].singlePN.animate"
   TextField "tfLablBtn02" at 215,50 size 40x25; Text '3'
      Visibility <- "Interface.btnRows[2].button.visibility"
      Appearance <- "Interface.btnRows[2].button.animate"
   TextField "tfAllottedBtn02" at 255,50 size 80x25; Text 'Text'
      Visibility <- "Interface.btnRows[2].total.visibility"
      Appearance <- "Interface.btnRows[2].total.animate"
   TextField "tfCriticalBtn02" at 335,50 size 80x25; Text 'Text'
      Visibility <- "Interface.btnRows[2].critical.visibility"
      Appearance <- "Interface.btnRows[2].critical.animate"
   TextField "tfPartNumberBtn02" at 415,50 size 256x25; Text 'Text'
      Visibility <- "Interface.btnRows[2].singlePN.visibility"
      Appearance <- "Interface.btnRows[2].singlePN.animate"
   TextField "tfLablBtn03" at 215,75 size 40x25; Text '4'
      Visibility <- "Interface.btnRows[3].button.visibility"
      Appearance <- "Interface.btnRows[3].button.animate"
   TextField "tfAllottedBtn03" at 255,75 size 80x25; Text 'Text'
      Visibility <- "Interface.btnRows[3].total.visibility"
      Appearance <- "Interface.btnRows[3].total.animate"
   TextField "tfCriticalBtn03" at 335,75 size 80x25; Text 'Text'
      Visibility <- "Interface.btnRows[3].critical.visibility"
      Appearance <- "Interface.btnRows[3].critical.animate"
   TextField "tfPartNumberBtn03" at 415,75 size 256x25; Text 'Text'
      Visibility <- "Interface.btnRows[3].singlePN.visibility"
      Appearance <- "Interface.btnRows[3].singlePN.animate"
   TextField "tfLablBtn04" at 215,100 size 40x25; Text '5'
      Visibility <- "Interface.btnRows[4].button.visibility"
      Appearance <- "Interface.btnRows[4].button.animate"
   TextField "tfAllottedBtn04" at 255,100 size 80x25; Text 'Text'
      Visibility <- "Interface.btnRows[4].total.visibility"
      Appearance <- "Interface.btnRows[4].total.animate"
   TextField "tfCriticalBtn04" at 335,100 size 80x25; Text 'Text'
      Visibility <- "Interface.btnRows[4].critical.visibility"
      Appearance <- "Interface.btnRows[4].critical.animate"
   TextField "tfPartNumberBtn04" at 415,100 size 256x25; Text 'Text'
      Visibility <- "Interface.btnRows[4].singlePN.visibility"
      Appearance <- "Interface.btnRows[4].singlePN.animate"
   TextField "tfLablBtn05" at 215,125 size 40x25; Text '6'
      Visibility <- "Interface.btnRows[5].button.visibility"
      Appearance <- "Interface.btnRows[5].button.animate"
   TextField "tfAllottedBtn05" at 255,125 size 80x25; Text 'Text'
      Visibility <- "Interface.btnRows[5].total.visibility"
      Appearance <- "Interface.btnRows[5].total.animate"
   TextField "tfCriticalBtn05" at 335,125 size 80x25; Text 'Text'
      Visibility <- "Interface.btnRows[5].critical.visibility"
      Appearance <- "Interface.btnRows[5].critical.animate"
   TextField "tfPartNumberBtn05" at 415,125 size 256x25; Text 'Text'
      Visibility <- "Interface.btnRows[5].singlePN.visibility"
      Appearance <- "Interface.btnRows[5].singlePN.animate"
   TextField "tfLablBtn06" at 215,150 size 40x25; Text '7'
      Visibility <- "Interface.btnRows[6].button.visibility"
      Appearance <- "Interface.btnRows[6].button.animate"
   TextField "tfAllottedBtn06" at 255,150 size 80x25; Text 'Text'
      Visibility <- "Interface.btnRows[6].total.visibility"
      Appearance <- "Interface.btnRows[6].total.animate"
   TextField "tfCriticalBtn06" at 335,150 size 80x25; Text 'Text'
      Visibility <- "Interface.btnRows[6].critical.visibility"
      Appearance <- "Interface.btnRows[6].critical.animate"
   TextField "tfPartNumberBtn06" at 415,150 size 256x25; Text 'Text'
      Visibility <- "Interface.btnRows[6].singlePN.visibility"
      Appearance <- "Interface.btnRows[6].singlePN.animate"
   TextField "tfLablBtn07" at 215,175 size 40x25; Text '8'
      Visibility <- "Interface.btnRows[7].button.visibility"
      Appearance <- "Interface.btnRows[7].button.animate"
   TextField "tfAllottedBtn07" at 255,175 size 80x25; Text 'Text'
      Visibility <- "Interface.btnRows[7].total.visibility"
      Appearance <- "Interface.btnRows[7].total.animate"
   TextField "tfCriticalBtn07" at 335,175 size 80x25; Text 'Text'
      Visibility <- "Interface.btnRows[7].critical.visibility"
      Appearance <- "Interface.btnRows[7].critical.animate"
   TextField "tfPartNumberBtn07" at 415,175 size 256x25; Text 'Text'
      Visibility <- "Interface.btnRows[7].singlePN.visibility"
      Appearance <- "Interface.btnRows[7].singlePN.animate"
   TextField "tfPNDoubleBtn00" at 415,0 size 256x25; Text 'Text'
      Visibility <- "Interface.btnRows[0].doublePN.visibility"
      Appearance <- "Interface.btnRows[0].doublePN.animate"
   TextField "tfPNDoubleBtn01" at 415,25 size 256x25; Text 'Text'
      Visibility <- "Interface.btnRows[1].doublePN.visibility"
      Appearance <- "Interface.btnRows[1].doublePN.animate"
   TextField "tfPNDoubleBtn02" at 415,50 size 256x25; Text 'Text'
      Visibility <- "Interface.btnRows[2].doublePN.visibility"
      Appearance <- "Interface.btnRows[2].doublePN.animate"
   TextField "tfPNDoubleBtn03" at 415,75 size 256x25; Text 'Text'
      Visibility <- "Interface.btnRows[3].doublePN.visibility"
      Appearance <- "Interface.btnRows[3].doublePN.animate"
   TextField "tfPNDoubleBtn04" at 415,100 size 256x25; Text 'Text'
      Visibility <- "Interface.btnRows[4].doublePN.visibility"
      Appearance <- "Interface.btnRows[4].doublePN.animate"
   TextField "tfPNDoubleBtn05" at 415,125 size 256x25; Text 'Text'
      Visibility <- "Interface.btnRows[5].doublePN.visibility"
      Appearance <- "Interface.btnRows[5].doublePN.animate"
   TextField "tfPNDoubleBtn06" at 415,150 size 256x25; Text 'Text'
      Visibility <- "Interface.btnRows[6].doublePN.visibility"
      Appearance <- "Interface.btnRows[6].doublePN.animate"
   TextField "tfPNDoubleBtn07" at 415,175 size 256x25; Text 'Text'
      Visibility <- "Interface.btnRows[7].doublePN.visibility"
      Appearance <- "Interface.btnRows[7].doublePN.animate"
*)

(* ===== HMI "HMI_RT_1" =====
system functions are stored by id; their names below are inferred from use

ScreenModuleEditorView "IO Field: Part Number: 2 Line" 370x111
   TextField "iofLabel2Line" at 0,0 size 235x37; Text 'Part Number:'
      Visibility <- "Interface.double_visible"
   Button "btnMode2Line" at 235,5 size 135x27; TextOff 'DOUBLE'
      on Press: function_b14e0dd5("Interface.double_actuate", 0)
      Visibility <- "Interface.double_visible"
      ObjectEnable <- "Interface.double_enable"
      Appearance <- "Interface.double_animate"
   IOField "iofPNTop" at 0,37 size 370x37; FormatPattern ????????????????????????????????????????
      on OnFinishInput: SetBit("Interface.double_input_finished_top")
      Visibility <- "Interface.double_visible"
      ProcessValue <- "Interface.double_value_top"
      ObjectEnable <- "Interface.double_enable"
   IOField "iofPNBottom" at 0,74 size 370x37; FormatPattern ????????????????????????????????????????
      on OnFinishInput: SetBit("Interface.double_input_finished_bottom")
      Visibility <- "Interface.double_visible"
      ProcessValue <- "Interface.double_value_bottom"
      ObjectEnable <- "Interface.double_enable"
   TextField "iofLabel1Line" at 0,0 size 235x55; Text 'Part Number:'
      Visibility <- "Interface.single_visible"
   Button "btnMode1Line" at 235,5 size 135x45; TextOff 'SINGLE'
      on Press: function_b14e0dd5("Interface.single_actuate", 0)
      Appearance <- "Interface.single_animate"
      ObjectEnable <- "Interface.single_enable"
      Visibility <- "Interface.single_visible"
   IOField "iofPN" at 0,55 size 370x56; FormatPattern ????????????????????????????????????????
      on OnFinishInput: SetBit("Interface.single_input_finished")
      Visibility <- "Interface.single_visible"
      ProcessValue <- "Interface.single_value"
      ObjectEnable <- "Interface.single_enable"
*)

(* ===== HMI "HMI_RT_1" =====
system functions are stored by id; their names below are inferred from use

ScreenModuleEditorView "IO Field: Part Number: 2 Line" 370x111
   TextField "iofLabel2Line" at 0,0 size 235x37; Text 'Part Number:'
      Visibility <- "Interface.double_visible"
   Button "btnMode2Line" at 235,5 size 135x27; TextOff 'DOUBLE'
      on Press: function_b14e0dd5("Interface.double_actuate", 0)
      Visibility <- "Interface.double_visible"
      ObjectEnable <- "Interface.double_enable"
      Appearance <- "Interface.double_animate"
   IOField "iofPNTop" at 0,37 size 370x34; FormatPattern ????????????????????????????????????????
      on OnFinishInput: SetBit("Interface.double_input_finished_top")
      Visibility <- "Interface.double_visible"
      ProcessValue <- "Interface.double_value_top"
      ObjectEnable <- "Interface.double_enable"
   IOField "iofPNBottom" at 0,77 size 370x34; FormatPattern ????????????????????????????????????????
      on OnFinishInput: SetBit("Interface.double_input_finished_bottom")
      Visibility <- "Interface.double_visible"
      ProcessValue <- "Interface.double_value_bottom"
      ObjectEnable <- "Interface.double_enable"
   TextField "iofLabel1Line" at 0,0 size 235x55; Text 'Part Number:'
      Visibility <- "Interface.single_visible"
   Button "btnMode1Line" at 235,5 size 135x45; TextOff 'SINGLE'
      on Press: function_b14e0dd5("Interface.single_actuate", 0)
      Appearance <- "Interface.single_animate"
      ObjectEnable <- "Interface.single_enable"
      Visibility <- "Interface.single_visible"
   IOField "iofPN" at 0,55 size 370x56; FormatPattern ????????????????????????????????????????
      on OnFinishInput: SetBit("Interface.single_input_finished")
      Visibility <- "Interface.single_visible"
      ProcessValue <- "Interface.single_value"
      ObjectEnable <- "Interface.single_enable"
*)

(* ===== HMI "HMI_RT_1" =====
system functions are stored by id; their names below are inferred from use

ScreenModuleEditorView "IO Field: Part Number: 2 Line" 370x111
   TextField "iofLabel2Line" at 0,0 size 235x37; Text 'Part Number:'
      Visibility <- "Interface.double_visible"
   Button "btnMode2Line" at 235,5 size 135x27; TextOff 'DOUBLE'
      on Press: function_b14e0dd5("Interface.double_actuate", 0)
      Visibility <- "Interface.double_visible"
      ObjectEnable <- "Interface.double_enable"
      Appearance <- "Interface.double_animate"
   IOField "iofPNTop" at 0,37 size 370x34; FormatPattern ????????????????????????????????????????
      on OnFinishInput: SetBit("Interface.double_input_finished_top")
      Visibility <- "Interface.double_visible"
      ProcessValue <- "Interface.double_value_top"
      ObjectEnable <- "Interface.double_enable"
   IOField "iofPNBottom" at 0,77 size 370x34; FormatPattern ????????????????????????????????????????
      on OnFinishInput: SetBit("Interface.double_input_finished_bottom")
      Visibility <- "Interface.double_visible"
      ProcessValue <- "Interface.double_value_bottom"
      ObjectEnable <- "Interface.double_enable"
   TextField "iofLabel1Line" at 0,0 size 235x55; Text 'Part Number:'
      Visibility <- "Interface.single_visible"
   Button "btnMode1Line" at 235,5 size 135x45; TextOff 'SINGLE'
      on Press: function_b14e0dd5("Interface.single_actuate", 0)
      Appearance <- "Interface.single_animate"
      ObjectEnable <- "Interface.single_enable"
      Visibility <- "Interface.single_visible"
   IOField "iofPN" at 0,55 size 370x56; FormatPattern ????????????????????????????????????????
      on OnFinishInput: SetBit("Interface.single_input_finished")
      Visibility <- "Interface.single_visible"
      ProcessValue <- "Interface.single_value"
      ObjectEnable <- "Interface.single_enable"
*)

(* ===== HMI "HMI_RT_1" =====

